screen "15卷绕经验参数" 1280x740, template "模板_调试"
   Group "Group_卷绕经验参数1" at 176,4 size 296x672; FormatPattern 99.99
   Group "Group_卷绕经验参数3" at 808,4 size 296x672; FormatPattern 99.99
   Group "Group_卷绕经验参数2" at 492,4 size 296x672; FormatPattern 99.99
   Button "OBJECT_3" at 176,4 size 80x38; TextOff '支数: / EXIT / 標準糸管１: / 표준보빈1:'
      on Press: SetTag("ST_HMI_Var_HMI_i16_Status_ShaGuan_Select", 1)
   Button "OBJECT_1" at 268,4 size 96x38; TextOff 'f1_n: / EXIT / 標準糸管１: / 표준보빈1:'
      on Press: SetTag("ST_HMI_Var_HMI_i16_Status_ShaGuan_Select", 1)
   Button "OBJECT_2" at 376,4 size 96x38; TextOff 'g1_n: / EXIT / 標準糸管１: / 표준보빈1:'
      on Press: SetTag("ST_HMI_Var_HMI_i16_Status_ShaGuan_Select", 1)
   IOField "IO Field_41" at 176,47 size 80x38; FormatPattern 99.9
      ProcessValue <- "ST_Calculation_Var_1_ZhiShu_ARRAY_JR{3}"
   IOField "IO Field_1" at 268,46 size 96x38; FormatPattern 99.999
      ProcessValue <- "ST_Calculation_Var_1_f1_n_delt_0_n_ARRAY_JR{3}"
   IOField "IO Field_2" at 376,46 size 96x38; FormatPattern 99.999
      ProcessValue <- "ST_Calculation_Var_1_g1_n_delt_0_n_ARRAY_JR{3}"
   IOField "IO Field_3" at 176,89 size 80x38; FormatPattern 99.9
      ProcessValue <- "ST_Calculation_Var_1_ZhiShu_ARRAY_JR{4}"
   IOField "IO Field_4" at 268,88 size 96x38; FormatPattern 99.999
      ProcessValue <- "ST_Calculation_Var_1_f1_n_delt_0_n_ARRAY_JR{4}"
   IOField "IO Field_5" at 376,88 size 96x38; FormatPattern 99.999
      ProcessValue <- "ST_Calculation_Var_1_g1_n_delt_0_n_ARRAY_JR{4}"
   IOField "IO Field_6" at 176,131 size 80x38; FormatPattern 99.9
      ProcessValue <- "ST_Calculation_Var_1_ZhiShu_ARRAY_JR{5}"
   IOField "IO Field_7" at 176,173 size 80x38; FormatPattern 99.9
      ProcessValue <- "ST_Calculation_Var_1_ZhiShu_ARRAY_JR{6}"
   IOField "IO Field_8" at 176,215 size 80x38; FormatPattern 99.9
      ProcessValue <- "ST_Calculation_Var_1_ZhiShu_ARRAY_JR{7}"
   IOField "IO Field_9" at 176,258 size 80x38; FormatPattern 99.9
      ProcessValue <- "ST_Calculation_Var_1_ZhiShu_ARRAY_JR{8}"
   IOField "IO Field_10" at 176,300 size 80x38; FormatPattern 99.9
      ProcessValue <- "ST_Calculation_Var_1_ZhiShu_ARRAY_JR{9}"
   IOField "IO Field_11" at 176,342 size 80x38; FormatPattern 99.9
      ProcessValue <- "ST_Calculation_Var_1_ZhiShu_ARRAY_JR{10}"
   IOField "IO Field_12" at 176,384 size 80x38; FormatPattern 99.9
      ProcessValue <- "ST_Calculation_Var_1_ZhiShu_ARRAY_JR{11}"
   IOField "IO Field_13" at 176,426 size 80x38; FormatPattern 99.9
      ProcessValue <- "ST_Calculation_Var_1_ZhiShu_ARRAY_JR{12}"
   IOField "IO Field_14" at 176,469 size 80x38; FormatPattern 99.9
      ProcessValue <- "ST_Calculation_Var_1_ZhiShu_ARRAY_JR{13}"
   IOField "IO Field_15" at 176,511 size 80x38; FormatPattern 99.9
      ProcessValue <- "ST_Calculation_Var_1_ZhiShu_ARRAY_JR{14}"
   IOField "IO Field_16" at 176,553 size 80x38; FormatPattern 99.9
      ProcessValue <- "ST_Calculation_Var_1_ZhiShu_ARRAY_JR{15}"
   IOField "IO Field_17" at 176,595 size 80x38; FormatPattern 99.9
      ProcessValue <- "ST_Calculation_Var_1_ZhiShu_ARRAY_JR{16}"
   IOField "IO Field_18" at 176,638 size 80x38; FormatPattern 99.9
      ProcessValue <- "ST_Calculation_Var_1_ZhiShu_ARRAY_JR{17}"
   IOField "IO Field_19" at 268,130 size 96x38; FormatPattern 99.999
      ProcessValue <- "ST_Calculation_Var_1_f1_n_delt_0_n_ARRAY_JR{5}"
   IOField "IO Field_20" at 268,172 size 96x38; FormatPattern 99.999
      ProcessValue <- "ST_Calculation_Var_1_f1_n_delt_0_n_ARRAY_JR{6}"
   IOField "IO Field_21" at 268,215 size 96x38; FormatPattern 99.999
      ProcessValue <- "ST_Calculation_Var_1_f1_n_delt_0_n_ARRAY_JR{7}"
   IOField "IO Field_22" at 268,257 size 96x38; FormatPattern 99.999
      ProcessValue <- "ST_Calculation_Var_1_f1_n_delt_0_n_ARRAY_JR{8}"
   IOField "IO Field_23" at 268,299 size 96x38; FormatPattern 99.999
      ProcessValue <- "ST_Calculation_Var_1_f1_n_delt_0_n_ARRAY_JR{9}"
   IOField "IO Field_24" at 268,342 size 96x38; FormatPattern 99.999
      ProcessValue <- "ST_Calculation_Var_1_f1_n_delt_0_n_ARRAY_JR{10}"
   IOField "IO Field_25" at 268,384 size 96x38; FormatPattern 99.999
      ProcessValue <- "ST_Calculation_Var_1_f1_n_delt_0_n_ARRAY_JR{11}"
   IOField "IO Field_26" at 268,426 size 96x38; FormatPattern 99.999
      ProcessValue <- "ST_Calculation_Var_1_f1_n_delt_0_n_ARRAY_JR{12}"
   IOField "IO Field_27" at 268,468 size 96x38; FormatPattern 99.999
      ProcessValue <- "ST_Calculation_Var_1_f1_n_delt_0_n_ARRAY_JR{13}"
   IOField "IO Field_28" at 268,511 size 96x38; FormatPattern 99.999
      ProcessValue <- "ST_Calculation_Var_1_f1_n_delt_0_n_ARRAY_JR{14}"
   IOField "IO Field_29" at 268,553 size 96x38; FormatPattern 99.999
      ProcessValue <- "ST_Calculation_Var_1_f1_n_delt_0_n_ARRAY_JR{15}"
   IOField "IO Field_30" at 268,595 size 96x38; FormatPattern 99.999
      ProcessValue <- "ST_Calculation_Var_1_f1_n_delt_0_n_ARRAY_JR{16}"
   IOField "IO Field_31" at 268,638 size 96x38; FormatPattern 99.999
      ProcessValue <- "ST_Calculation_Var_1_f1_n_delt_0_n_ARRAY_JR{17}"
   IOField "IO Field_32" at 376,130 size 96x38; FormatPattern 99.999
      ProcessValue <- "ST_Calculation_Var_1_g1_n_delt_0_n_ARRAY_JR{5}"
   IOField "IO Field_33" at 376,172 size 96x38; FormatPattern 99.999
      ProcessValue <- "ST_Calculation_Var_1_g1_n_delt_0_n_ARRAY_JR{6}"
   IOField "IO Field_34" at 376,215 size 96x38; FormatPattern 99.999
      ProcessValue <- "ST_Calculation_Var_1_g1_n_delt_0_n_ARRAY_JR{7}"
   IOField "IO Field_35" at 376,257 size 96x38; FormatPattern 99.999
      ProcessValue <- "ST_Calculation_Var_1_g1_n_delt_0_n_ARRAY_JR{8}"
   IOField "IO Field_36" at 376,299 size 96x38; FormatPattern 99.999
      ProcessValue <- "ST_Calculation_Var_1_g1_n_delt_0_n_ARRAY_JR{9}"
   IOField "IO Field_37" at 376,342 size 96x38; FormatPattern 99.999
      ProcessValue <- "ST_Calculation_Var_1_g1_n_delt_0_n_ARRAY_JR{10}"
   IOField "IO Field_38" at 376,384 size 96x38; FormatPattern 99.999
      ProcessValue <- "ST_Calculation_Var_1_g1_n_delt_0_n_ARRAY_JR{11}"
   IOField "IO Field_39" at 376,426 size 96x38; FormatPattern 99.999
      ProcessValue <- "ST_Calculation_Var_1_g1_n_delt_0_n_ARRAY_JR{12}"
   IOField "IO Field_40" at 376,468 size 96x38; FormatPattern 99.999
      ProcessValue <- "ST_Calculation_Var_1_g1_n_delt_0_n_ARRAY_JR{13}"
   IOField "IO Field_42" at 376,511 size 96x38; FormatPattern 99.999
      ProcessValue <- "ST_Calculation_Var_1_g1_n_delt_0_n_ARRAY_JR{14}"
   IOField "IO Field_43" at 376,553 size 96x38; FormatPattern 99.999
      ProcessValue <- "ST_Calculation_Var_1_g1_n_delt_0_n_ARRAY_JR{15}"
   IOField "IO Field_44" at 376,595 size 96x38; FormatPattern 99.999
      ProcessValue <- "ST_Calculation_Var_1_g1_n_delt_0_n_ARRAY_JR{16}"
   IOField "IO Field_45" at 376,638 size 96x38; FormatPattern 99.999
      ProcessValue <- "ST_Calculation_Var_1_g1_n_delt_0_n_ARRAY_JR{17}"
   Button "OBJECT_7" at 808,4 size 80x38; TextOff '支数: / EXIT / 標準糸管１: / 표준보빈1:'
      on Press: SetTag("ST_HMI_Var_HMI_i16_Status_ShaGuan_Select", 1)
   Button "OBJECT_8" at 900,4 size 96x38; TextOff 'f1_n: / EXIT / 標準糸管１: / 표준보빈1:'
      on Press: SetTag("ST_HMI_Var_HMI_i16_Status_ShaGuan_Select", 1)
   Button "OBJECT_9" at 1008,4 size 96x38; TextOff 'g1_n: / EXIT / 標準糸管１: / 표준보빈1:'
      on Press: SetTag("ST_HMI_Var_HMI_i16_Status_ShaGuan_Select", 1)
   IOField "IO Field_91" at 808,47 size 80x38; FormatPattern 99.9
      ProcessValue <- "ST_Calculation_Var_1_ZhiShu_ARRAY_JR{33}"
   IOField "IO Field_92" at 900,46 size 96x38; FormatPattern 99.999
      ProcessValue <- "ST_Calculation_Var_1_f1_n_delt_0_n_ARRAY_JR{33}"
   IOField "IO Field_93" at 1008,46 size 96x38; FormatPattern 99.999
      ProcessValue <- "ST_Calculation_Var_1_g1_n_delt_0_n_ARRAY_JR{33}"
   IOField "IO Field_94" at 808,89 size 80x38; FormatPattern 99.9
      ProcessValue <- "ST_Calculation_Var_1_ZhiShu_ARRAY_JR{34}"
   IOField "IO Field_95" at 900,88 size 96x38; FormatPattern 99.999
      ProcessValue <- "ST_Calculation_Var_1_f1_n_delt_0_n_ARRAY_JR{34}"
   IOField "IO Field_96" at 1008,88 size 96x38; FormatPattern 99.999
      ProcessValue <- "ST_Calculation_Var_1_g1_n_delt_0_n_ARRAY_JR{34}"
   IOField "IO Field_97" at 808,131 size 80x38; FormatPattern 99.9
      ProcessValue <- "ST_Calculation_Var_1_ZhiShu_ARRAY_JR{35}"
   IOField "IO Field_98" at 808,173 size 80x38; FormatPattern 99.9
      ProcessValue <- "ST_Calculation_Var_1_ZhiShu_ARRAY_JR{36}"
   IOField "IO Field_99" at 808,215 size 80x38; FormatPattern 99.9
      ProcessValue <- "ST_Calculation_Var_1_ZhiShu_ARRAY_JR{37}"
   IOField "IO Field_100" at 808,258 size 80x38; FormatPattern 99.9
      ProcessValue <- "ST_Calculation_Var_1_ZhiShu_ARRAY_JR{38}"
   IOField "IO Field_101" at 808,300 size 80x38; FormatPattern 99.9
      ProcessValue <- "ST_Calculation_Var_1_ZhiShu_ARRAY_JR{39}"
   IOField "IO Field_102" at 808,342 size 80x38; FormatPattern 99.9
      ProcessValue <- "ST_Calculation_Var_1_ZhiShu_ARRAY_JR{40}"
   IOField "IO Field_103" at 808,384 size 80x38; FormatPattern 99.9
      ProcessValue <- "ST_Calculation_Var_1_ZhiShu_ARRAY_JR{41}"
   IOField "IO Field_104" at 808,426 size 80x38; FormatPattern 99.9
      ProcessValue <- "ST_Calculation_Var_1_ZhiShu_ARRAY_JR{42}"
   IOField "IO Field_105" at 808,469 size 80x38; FormatPattern 99.9
      ProcessValue <- "ST_Calculation_Var_1_ZhiShu_ARRAY_JR{43}"
   IOField "IO Field_106" at 808,511 size 80x38; FormatPattern 99.9
      ProcessValue <- "ST_Calculation_Var_1_ZhiShu_ARRAY_JR{44}"
   IOField "IO Field_107" at 808,553 size 80x38; FormatPattern 99.9
      ProcessValue <- "ST_Calculation_Var_1_ZhiShu_ARRAY_JR{45}"
   IOField "IO Field_108" at 808,595 size 80x38; FormatPattern 99.9
      ProcessValue <- "ST_Calculation_Var_1_ZhiShu_ARRAY_JR{46}"
   IOField "IO Field_109" at 808,638 size 80x38; FormatPattern 99.9
      ProcessValue <- "ST_Calculation_Var_1_ZhiShu_ARRAY_JR{47}"
   IOField "IO Field_110" at 900,130 size 96x38; FormatPattern 99.999
      ProcessValue <- "ST_Calculation_Var_1_f1_n_delt_0_n_ARRAY_JR{35}"
   IOField "IO Field_111" at 900,172 size 96x38; FormatPattern 99.999
      ProcessValue <- "ST_Calculation_Var_1_f1_n_delt_0_n_ARRAY_JR{36}"
   IOField "IO Field_112" at 900,215 size 96x38; FormatPattern 99.999
      ProcessValue <- "ST_Calculation_Var_1_f1_n_delt_0_n_ARRAY_JR{37}"
   IOField "IO Field_113" at 900,257 size 96x38; FormatPattern 99.999
      ProcessValue <- "ST_Calculation_Var_1_f1_n_delt_0_n_ARRAY_JR{38}"
   IOField "IO Field_114" at 900,299 size 96x38; FormatPattern 99.999
      ProcessValue <- "ST_Calculation_Var_1_f1_n_delt_0_n_ARRAY_JR{39}"
   IOField "IO Field_115" at 900,342 size 96x38; FormatPattern 99.999
      ProcessValue <- "ST_Calculation_Var_1_f1_n_delt_0_n_ARRAY_JR{40}"
   IOField "IO Field_116" at 900,384 size 96x38; FormatPattern 99.999
      ProcessValue <- "ST_Calculation_Var_1_f1_n_delt_0_n_ARRAY_JR{41}"
   IOField "IO Field_117" at 900,426 size 96x38; FormatPattern 99.999
      ProcessValue <- "ST_Calculation_Var_1_f1_n_delt_0_n_ARRAY_JR{42}"
   IOField "IO Field_118" at 900,468 size 96x38; FormatPattern 99.999
      ProcessValue <- "ST_Calculation_Var_1_f1_n_delt_0_n_ARRAY_JR{43}"
   IOField "IO Field_119" at 900,511 size 96x38; FormatPattern 99.999
      ProcessValue <- "ST_Calculation_Var_1_f1_n_delt_0_n_ARRAY_JR{44}"
   IOField "IO Field_120" at 900,553 size 96x38; FormatPattern 99.999
      ProcessValue <- "ST_Calculation_Var_1_f1_n_delt_0_n_ARRAY_JR{45}"
   IOField "IO Field_121" at 900,595 size 96x38; FormatPattern 99.999
      ProcessValue <- "ST_Calculation_Var_1_f1_n_delt_0_n_ARRAY_JR{46}"
   IOField "IO Field_122" at 900,638 size 96x38; FormatPattern 99.999
      ProcessValue <- "ST_Calculation_Var_1_f1_n_delt_0_n_ARRAY_JR{47}"
   IOField "IO Field_123" at 1008,130 size 96x38; FormatPattern 99.999
      ProcessValue <- "ST_Calculation_Var_1_g1_n_delt_0_n_ARRAY_JR{35}"
   IOField "IO Field_124" at 1008,172 size 96x38; FormatPattern 99.999
      ProcessValue <- "ST_Calculation_Var_1_g1_n_delt_0_n_ARRAY_JR{36}"
   IOField "IO Field_125" at 1008,215 size 96x38; FormatPattern 99.999
      ProcessValue <- "ST_Calculation_Var_1_g1_n_delt_0_n_ARRAY_JR{37}"
   IOField "IO Field_126" at 1008,257 size 96x38; FormatPattern 99.999
      ProcessValue <- "ST_Calculation_Var_1_g1_n_delt_0_n_ARRAY_JR{38}"
   IOField "IO Field_127" at 1008,299 size 96x38; FormatPattern 99.999
      ProcessValue <- "ST_Calculation_Var_1_g1_n_delt_0_n_ARRAY_JR{39}"
   IOField "IO Field_128" at 1008,342 size 96x38; FormatPattern 99.999
      ProcessValue <- "ST_Calculation_Var_1_g1_n_delt_0_n_ARRAY_JR{40}"
   IOField "IO Field_129" at 1008,384 size 96x38; FormatPattern 99.999
      ProcessValue <- "ST_Calculation_Var_1_g1_n_delt_0_n_ARRAY_JR{41}"
   IOField "IO Field_130" at 1008,426 size 96x38; FormatPattern 99.999
      ProcessValue <- "ST_Calculation_Var_1_g1_n_delt_0_n_ARRAY_JR{42}"
   IOField "IO Field_131" at 1008,468 size 96x38; FormatPattern 99.999
      ProcessValue <- "ST_Calculation_Var_1_g1_n_delt_0_n_ARRAY_JR{43}"
   IOField "IO Field_132" at 1008,511 size 96x38; FormatPattern 99.999
      ProcessValue <- "ST_Calculation_Var_1_g1_n_delt_0_n_ARRAY_JR{44}"
   IOField "IO Field_133" at 1008,553 size 96x38; FormatPattern 99.999
      ProcessValue <- "ST_Calculation_Var_1_g1_n_delt_0_n_ARRAY_JR{45}"
   IOField "IO Field_134" at 1008,595 size 96x38; FormatPattern 99.999
      ProcessValue <- "ST_Calculation_Var_1_g1_n_delt_0_n_ARRAY_JR{46}"
   IOField "IO Field_135" at 1008,638 size 96x38; FormatPattern 99.999
      ProcessValue <- "ST_Calculation_Var_1_g1_n_delt_0_n_ARRAY_JR{47}"
   Button "OBJECT_4" at 492,4 size 80x38; TextOff '支数: / EXIT / 標準糸管１: / 표준보빈1:'
      on Press: SetTag("ST_HMI_Var_HMI_i16_Status_ShaGuan_Select", 1)
   Button "OBJECT_5" at 584,4 size 96x38; TextOff 'f1_n: / EXIT / 標準糸管１: / 표준보빈1:'
      on Press: SetTag("ST_HMI_Var_HMI_i16_Status_ShaGuan_Select", 1)
   Button "OBJECT_6" at 692,4 size 96x38; TextOff 'g1_n: / EXIT / 標準糸管１: / 표준보빈1:'
      on Press: SetTag("ST_HMI_Var_HMI_i16_Status_ShaGuan_Select", 1)
   IOField "IO Field_46" at 492,47 size 80x38; FormatPattern 99.9
      ProcessValue <- "ST_Calculation_Var_1_ZhiShu_ARRAY_JR{18}"
   IOField "IO Field_47" at 584,46 size 96x38; FormatPattern 99.999
      ProcessValue <- "ST_Calculation_Var_1_f1_n_delt_0_n_ARRAY_JR{18}"
   IOField "IO Field_48" at 692,46 size 96x38; FormatPattern 99.999
      ProcessValue <- "ST_Calculation_Var_1_g1_n_delt_0_n_ARRAY_JR{18}"
   IOField "IO Field_49" at 492,89 size 80x38; FormatPattern 99.9
      ProcessValue <- "ST_Calculation_Var_1_ZhiShu_ARRAY_JR{19}"
   IOField "IO Field_50" at 584,88 size 96x38; FormatPattern 99.999
      ProcessValue <- "ST_Calculation_Var_1_f1_n_delt_0_n_ARRAY_JR{19}"
   IOField "IO Field_51" at 692,88 size 96x38; FormatPattern 99.999
      ProcessValue <- "ST_Calculation_Var_1_g1_n_delt_0_n_ARRAY_JR{19}"
   IOField "IO Field_52" at 492,131 size 80x38; FormatPattern 99.9
      ProcessValue <- "ST_Calculation_Var_1_ZhiShu_ARRAY_JR{20}"
   IOField "IO Field_53" at 492,173 size 80x38; FormatPattern 99.9
      ProcessValue <- "ST_Calculation_Var_1_ZhiShu_ARRAY_JR{21}"
   IOField "IO Field_54" at 492,215 size 80x38; FormatPattern 99.9
      ProcessValue <- "ST_Calculation_Var_1_ZhiShu_ARRAY_JR{22}"
   IOField "IO Field_55" at 492,258 size 80x38; FormatPattern 99.9
      ProcessValue <- "ST_Calculation_Var_1_ZhiShu_ARRAY_JR{23}"
   IOField "IO Field_56" at 492,300 size 80x38; FormatPattern 99.9
      ProcessValue <- "ST_Calculation_Var_1_ZhiShu_ARRAY_JR{24}"
   IOField "IO Field_57" at 492,342 size 80x38; FormatPattern 99.9
      ProcessValue <- "ST_Calculation_Var_1_ZhiShu_ARRAY_JR{25}"
   IOField "IO Field_58" at 492,384 size 80x38; FormatPattern 99.9
      ProcessValue <- "ST_Calculation_Var_1_ZhiShu_ARRAY_JR{26}"
   IOField "IO Field_59" at 492,426 size 80x38; FormatPattern 99.9
      ProcessValue <- "ST_Calculation_Var_1_ZhiShu_ARRAY_JR{27}"
   IOField "IO Field_60" at 492,469 size 80x38; FormatPattern 99.9
      ProcessValue <- "ST_Calculation_Var_1_ZhiShu_ARRAY_JR{28}"
   IOField "IO Field_61" at 492,511 size 80x38; FormatPattern 99.9
      ProcessValue <- "ST_Calculation_Var_1_ZhiShu_ARRAY_JR{29}"
   IOField "IO Field_62" at 492,553 size 80x38; FormatPattern 99.9
      ProcessValue <- "ST_Calculation_Var_1_ZhiShu_ARRAY_JR{30}"
   IOField "IO Field_63" at 492,595 size 80x38; FormatPattern 99.9
      ProcessValue <- "ST_Calculation_Var_1_ZhiShu_ARRAY_JR{31}"
   IOField "IO Field_64" at 492,638 size 80x38; FormatPattern 99.9
      ProcessValue <- "ST_Calculation_Var_1_ZhiShu_ARRAY_JR{32}"
   IOField "IO Field_65" at 584,130 size 96x38; FormatPattern 99.999
      ProcessValue <- "ST_Calculation_Var_1_f1_n_delt_0_n_ARRAY_JR{20}"
   IOField "IO Field_66" at 584,172 size 96x38; FormatPattern 99.999
      ProcessValue <- "ST_Calculation_Var_1_f1_n_delt_0_n_ARRAY_JR{21}"
   IOField "IO Field_67" at 584,215 size 96x38; FormatPattern 99.999
      ProcessValue <- "ST_Calculation_Var_1_f1_n_delt_0_n_ARRAY_JR{22}"
   IOField "IO Field_68" at 584,257 size 96x38; FormatPattern 99.999
      ProcessValue <- "ST_Calculation_Var_1_f1_n_delt_0_n_ARRAY_JR{23}"
   IOField "IO Field_69" at 584,299 size 96x38; FormatPattern 99.999
      ProcessValue <- "ST_Calculation_Var_1_f1_n_delt_0_n_ARRAY_JR{24}"
   IOField "IO Field_70" at 584,342 size 96x38; FormatPattern 99.999
      ProcessValue <- "ST_Calculation_Var_1_f1_n_delt_0_n_ARRAY_JR{25}"
   IOField "IO Field_71" at 584,384 size 96x38; FormatPattern 99.999
      ProcessValue <- "ST_Calculation_Var_1_f1_n_delt_0_n_ARRAY_JR{26}"
   IOField "IO Field_72" at 584,426 size 96x38; FormatPattern 99.999
      ProcessValue <- "ST_Calculation_Var_1_f1_n_delt_0_n_ARRAY_JR{27}"
   IOField "IO Field_73" at 584,468 size 96x38; FormatPattern 99.999
      ProcessValue <- "ST_Calculation_Var_1_f1_n_delt_0_n_ARRAY_JR{28}"
   IOField "IO Field_74" at 584,511 size 96x38; FormatPattern 99.999
      ProcessValue <- "ST_Calculation_Var_1_f1_n_delt_0_n_ARRAY_JR{29}"
   IOField "IO Field_75" at 584,553 size 96x38; FormatPattern 99.999
      ProcessValue <- "ST_Calculation_Var_1_f1_n_delt_0_n_ARRAY_JR{30}"
   IOField "IO Field_76" at 584,595 size 96x38; FormatPattern 99.999
      ProcessValue <- "ST_Calculation_Var_1_f1_n_delt_0_n_ARRAY_JR{31}"
   IOField "IO Field_77" at 584,638 size 96x38; FormatPattern 99.999
      ProcessValue <- "ST_Calculation_Var_1_f1_n_delt_0_n_ARRAY_JR{32}"
   IOField "IO Field_78" at 692,130 size 96x38; FormatPattern 99.999
      ProcessValue <- "ST_Calculation_Var_1_g1_n_delt_0_n_ARRAY_JR{20}"
   IOField "IO Field_79" at 692,172 size 96x38; FormatPattern 99.999
      ProcessValue <- "ST_Calculation_Var_1_g1_n_delt_0_n_ARRAY_JR{21}"
   IOField "IO Field_80" at 692,215 size 96x38; FormatPattern 99.999
      ProcessValue <- "ST_Calculation_Var_1_g1_n_delt_0_n_ARRAY_JR{22}"
   IOField "IO Field_81" at 692,257 size 96x38; FormatPattern 99.999
      ProcessValue <- "ST_Calculation_Var_1_g1_n_delt_0_n_ARRAY_JR{23}"
   IOField "IO Field_82" at 692,299 size 96x38; FormatPattern 99.999
      ProcessValue <- "ST_Calculation_Var_1_g1_n_delt_0_n_ARRAY_JR{24}"
   IOField "IO Field_83" at 692,342 size 96x38; FormatPattern 99.999
      ProcessValue <- "ST_Calculation_Var_1_g1_n_delt_0_n_ARRAY_JR{25}"
   IOField "IO Field_84" at 692,384 size 96x38; FormatPattern 99.999
      ProcessValue <- "ST_Calculation_Var_1_g1_n_delt_0_n_ARRAY_JR{26}"
   IOField "IO Field_85" at 692,426 size 96x38; FormatPattern 99.999
      ProcessValue <- "ST_Calculation_Var_1_g1_n_delt_0_n_ARRAY_JR{27}"
   IOField "IO Field_86" at 692,468 size 96x38; FormatPattern 99.999
      ProcessValue <- "ST_Calculation_Var_1_g1_n_delt_0_n_ARRAY_JR{28}"
   IOField "IO Field_87" at 692,511 size 96x38; FormatPattern 99.999
      ProcessValue <- "ST_Calculation_Var_1_g1_n_delt_0_n_ARRAY_JR{29}"
   IOField "IO Field_88" at 692,553 size 96x38; FormatPattern 99.999
      ProcessValue <- "ST_Calculation_Var_1_g1_n_delt_0_n_ARRAY_JR{30}"
   IOField "IO Field_89" at 692,595 size 96x38; FormatPattern 99.999
      ProcessValue <- "ST_Calculation_Var_1_g1_n_delt_0_n_ARRAY_JR{31}"
   IOField "IO Field_90" at 692,638 size 96x38; FormatPattern 99.999
      ProcessValue <- "ST_Calculation_Var_1_g1_n_delt_0_n_ARRAY_JR{32}"

screen "16机械参数" 1280x740, template "模板_调试"
   GraphicView "图形视图_1" at 395,6 size 437x668; Picture "成形参数_400×600"
   TextField "文本域_1" at 847,6 size 298x260; Text '测绘尺寸: rc0 :成形弓半径 rz0 :张力弓半径 xco :成形弓圆心x坐标 yco :成形弓圆心y坐标 hcz :轴心高度差 H :锭子总高度 Dl :罗拉直径 Hld :锭尖到罗拉顶部的高度 Lld :锭尖到罗拉的距离'
   TextField "文本域_3" at 847,355 size 298x250; Text '绘图后得出的： xzo :张力弓圆心x坐标 yzo :张力弓圆心y坐标 xit_0 :成形弓零位对应的角度 GAM_max :张力弓零位对应的角度 xit_delt_max :成形弓最大行程 gam_delt_max :张力弓最大行程 X_L_0 :罗拉最高点x坐标 Y_L_0 :罗拉最高点y坐标'
   TextField "文本域_2" at 847,270 size 298x80; Text '调整尺寸： hc0 :成形弓零位到锭尖的高度 hz0 :张力弓零位到锭尖的高度'
   TextField "文本域_4" at 143,22 size 145x30; Text '1.rc0'
   TextField "文本域_5" at 143,77 size 145x30; Text '2.rz0'
   TextField "文本域_6" at 143,132 size 145x30; Text '3.xco'
   TextField "文本域_7" at 143,187 size 145x30; Text '4.yco'
   TextField "文本域_8" at 143,242 size 145x30; Text '5.xzo'
   TextField "文本域_9" at 143,297 size 145x30; Text '6.yzo'
   TextField "文本域_10" at 143,352 size 145x30; Text '7.xit_0'
   TextField "文本域_11" at 143,407 size 145x30; Text '8.GAM_max'
   TextField "文本域_12" at 143,462 size 145x30; Text '9.xit_delt_max'
   TextField "文本域_13" at 143,517 size 145x30; Text '10.X_L_0'
   TextField "文本域_14" at 143,572 size 145x30; Text '11.Y_L_0'
   TextField "文本域_15" at 143,628 size 145x30; Text '12.CX_max'
   TextField "文本域_16" at 847,610 size 298x63; Text '设定参数： CX_max :落纱成形最低位置'
   IOField "IO Field_9" at 304,22 size 80x30
      ProcessValue <- "ST_HMI_Var_HMI_rc0"
   IOField "IO Field_1" at 304,77 size 80x30
      ProcessValue <- "ST_HMI_Var_HMI_rz0"
   IOField "IO Field_2" at 304,132 size 80x30
      ProcessValue <- "ST_HMI_Var_HMI_xco"
   IOField "IO Field_3" at 304,187 size 80x30
      ProcessValue <- "ST_HMI_Var_HMI_yco"
   IOField "IO Field_4" at 304,242 size 80x30
      ProcessValue <- "ST_HMI_Var_HMI_xzo"
   IOField "IO Field_5" at 304,297 size 80x30
      ProcessValue <- "ST_HMI_Var_HMI_yzo"
   IOField "IO Field_6" at 304,352 size 80x30
      ProcessValue <- "ST_HMI_Var_HMI_xit_0"
   IOField "IO Field_7" at 304,407 size 80x30
      ProcessValue <- "ST_HMI_Var_HMI_GAM_max"
   IOField "IO Field_8" at 304,462 size 80x30
      ProcessValue <- "ST_HMI_Var_HMI_xit_delt_max"
   IOField "IO Field_10" at 304,517 size 80x30
      ProcessValue <- "ST_HMI_Var_HMI_X_L_0"
   IOField "IO Field_11" at 304,572 size 80x30
      ProcessValue <- "ST_HMI_Var_HMI_Y_L_0"
   IOField "IO Field_12" at 304,628 size 80x30
      ProcessValue <- "ST_HMI_Var_HMI_r64Position_ChengXing_Botton"

Template "模板_根" 1280x740
   Button "template_1_1" at 80,680 size 80x60; TextOn '手动画面'; TextOff '手动操作'; PictureOn "manual_5_500×500_反相"; PictureOff "manual_5_500×500"
      on Release: ActivateScreenByNumber("Picture", 0)
      on Press: SetTag("Picture", 5)
      Appearance <- "Picture"
   Button "template_1_2" at 720,680 size 80x60; TextOn '报警画面'; TextOff '报 警'; PictureOn "emblem_important_1_200×200_反相"; PictureOff "emblem_important_1_200×200"
      on Release: ActivateScreenByNumber("Picture", 0)
      on Press: SetTag("Picture", 6)
      Appearance <- "Picture"
   Button "template_1_5" at 800,680 size 80x60; TextOn '保养提示'; TextOff '保养提示'; PictureOn "baoyang_6_600×600_反相"; PictureOff "baoyang_6_600×600"
      on Release: ActivateScreenByNumber("Picture", 0)
      on Press: SetTag("Picture", 8)
      Appearance <- "Picture"
   Button "template_1_7" at 880,680 size 80x60; TextOn '调试画面'; TextOff '调 试'; Authorization "Operate_4"; PictureOff "kdeconnect-tray_100×100"; PictureOn "kdeconnect-tray_100×100_反相"
      on Release: ActivateScreenByNumber("Picture", 0); function_f23ef4c9()
      on Press: SetTag("Picture", 3)
      Appearance <- "Picture"
   Button "template_1_3" at 0,680 size 80x60; TextOn '手动画面'; TextOff '手动操作'; PictureOff "图形_16"
      on Release: ActivateScreenByNumber("Picture", 0); SetTag("ST_HMI_Var_HMI_i32_ZouChe_ZhanJu_ss_1", 0)
      on Press: function_f23ef4c9(); SetTag("Picture", 1)
      Appearance <- "Picture"
   Button "template_1_4" at 1120,680 size 80x60; TextOff '调 试'; TextOn '调试画面'; Authorization "Operate_4"; PictureOff "System_Shutdown_100×100"; PictureOn "System_Shutdown_反相_100×100"
      on Click: function_f23ef4c9()
      on Release: StopRuntime(0)
   Button "template_1_6" at 1040,680 size 80x60; TextOff 'Text'; TextOn '调试画面'; Authorization "Operate_4"; PictureOff "computer_laptop_100×100"; PictureOn "computer_laptop_100×100_反相"
      on Click: function_f23ef4c9()
      on Release: function_f34a74f3()
   Button "template_1_8" at 960,680 size 80x60; TextOff 'Text'; TextOn '调试画面'; Authorization "Operate_4"; PictureOff "similarartists_amarok_100×100"; PictureOn "similarartists_amarok_100×100_反相"
      on Release: ActivateScreenByNumber("Picture", 0)
      on Press: SetTag("Picture", 7)
      Appearance <- "Picture"
   Button "template_1_23" at 160,680 size 160x60; TextOn '工艺'; TextOff '工艺'; PictureOn "settings_1_32×32_反相"; PictureOff "settings_1_32×32"
      on Release: ActivateScreenByNumber("Picture", 0)
      on Press: SetTag("Picture", 2)
      Appearance <- "Picture"
   TextField "模板_文本域_2" at 320,680 size 400x60; Text '苏州友联纺工装备科技股份有限公司'
   Button "OBJECT_122" at 1200,680 size 80x60; TextOn '响 铃'; TextOff '响 铃 / EXIT'; PictureOn "Gold_bell_100×100_反相"; PictureOff "Gold_bell_100×100"
      on Release: ResetBit("ST_HMI_Var_HMI_bo_XiangLing")
      on Press: SetBit("ST_HMI_Var_HMI_bo_XiangLing")
      Appearance <- "ST_HMI_Var_HMI_bo_XiangLing"

Template "模板_动画" 1280x740
   Bar "棒图_2" at 116,16 size 17x416; MinimumValue -1000; MaximumValue 10500
      ProcessValue <- "ST_HMI_Var_HMI_r64Axis_DingZi_Velocity_real"
   Group "Group_锭子转速" at 163,92 size 84x50
   Group "Group_动画_1" at 160,100 size 1103x448
   Group "Group_捻度" at 163,155 size 98x50
   Button "template_animation_1" at 80,680 size 80x60; TextOn '手动画面'; TextOff '手动操作'; PictureOn "manual_5_500×500_反相"; PictureOff "manual_5_500×500"
      on Release: ActivateScreenByNumber("Picture", 0)
      on Press: SetTag("Picture", 5)
      Appearance <- "Picture"
   Button "template_animation_2" at 720,680 size 80x60; TextOn '报警画面'; TextOff '报 警'; PictureOn "emblem_important_1_200×200_反相"; PictureOff "emblem_important_1_200×200"
      on Release: ActivateScreenByNumber("Picture", 0)
      on Press: SetTag("Picture", 6)
      Appearance <- "Picture"
   Button "template_animation_5" at 800,680 size 80x60; TextOn '保养提示'; TextOff '保养提示'; PictureOn "baoyang_6_600×600_反相"; PictureOff "baoyang_6_600×600"
      on Release: ActivateScreenByNumber("Picture", 0)
      on Press: SetTag("Picture", 8)
      Appearance <- "Picture"
   Button "template_animation_7" at 880,680 size 80x60; TextOn '调试画面'; TextOff '调 试'; Authorization "Operate_4"; PictureOff "kdeconnect-tray_100×100"; PictureOn "kdeconnect-tray_100×100_反相"
      on Release: ActivateScreenByNumber("Picture", 0); function_f23ef4c9()
      on Press: SetTag("Picture", 3)
      Appearance <- "Picture"
   Button "template_animation_3" at 0,680 size 80x60; TextOn '手动画面'; TextOff '手动操作'; PictureOff "图形_16"
      on Release: ActivateScreenByNumber("Picture", 0); SetTag("ST_HMI_Var_HMI_i32_ZouChe_ZhanJu_ss_1", 0)
      on Press: function_f23ef4c9(); SetTag("Picture", 1)
      Appearance <- "Picture"
   Button "template_animation_4" at 1120,680 size 80x60; TextOff '调 试'; TextOn '调试画面'; PictureOn "System_Shutdown_反相_100×100"; PictureOff "System_Shutdown_100×100"; Authorization "Operate_4"
      on Click: function_f23ef4c9()
      on Release: StopRuntime(0)
   Button "template_animation_6" at 1040,680 size 80x60; TextOff 'Text'; TextOn '调试画面'; PictureOn "computer_laptop_100×100_反相"; PictureOff "computer_laptop_100×100"; Authorization "Operate_4"
      on Click: function_f23ef4c9()
      on Release: function_f34a74f3()
   Button "template_animation_8" at 960,680 size 80x60; TextOff 'Text'; TextOn '调试画面'; PictureOn "similarartists_amarok_100×100_反相"; PictureOff "similarartists_amarok_100×100"; Authorization "Operate_4"
      on Release: ActivateScreenByNumber("Picture", 0)
      on Press: SetTag("Picture", 7)
      Appearance <- "Picture"
   Rectangle "模板_矩形_2" at 559,499 size 552x50
      Visibility <- "ST_Main_Var_g_bo_Automatic_Running_Status"
   Button "template_animation_23" at 160,680 size 160x60; TextOn '工艺'; TextOff '工艺'; PictureOn "settings_1_32×32_反相"; PictureOff "settings_1_32×32"
      on Release: ActivateScreenByNumber("Picture", 0)
      on Press: SetTag("Picture", 2)
      Appearance <- "Picture"
   TextField "模板_文本域_2" at 320,680 size 400x60; Text '苏州友联纺工装备科技股份有限公司'
   IOField "IO Field_57" at 163,92 size 51x25; FormatPattern 99999
      ProcessValue <- "ST_HMI_Var_HMI_r64Axis_DingZi_Velocity_real"
   TextField "文本域_9" at 213,92 size 34x25; Text '/'
   IOField "IO Field_56" at 163,117 size 51x25; FormatPattern 99999
      ProcessValue <- "ST_HMI_Var_HMI_r64Axis_DingZi_Velocity_object"
   TextField "文本域_10" at 213,117 size 34x25; Text 'rpm'
   Group "Group_纱穗" at 11,16 size 78x416
   Polygon "多边形_195" at 11,122 size 78x280
      Visibility <- "VBS_hengsi_status1"
   Polygon "多边形_196" at 11,207 size 78x195
      Visibility <- "VBS_hengsi_status1"
   Polygon "多边形_264" at 32,301 size 38x101
      Visibility <- "VBS_hengsi_status0"
   Polygon "多边形_265" at 36,312 size 29x90
      Visibility <- "VBS_hengsi_status0"
   Polygon "多边形_198" at 11,116 size 78x286
      Visibility <- "VBS_hengsi_status1"
   Polygon "多边形_199" at 11,201 size 78x200
      Visibility <- "VBS_hengsi_status1"
   Polygon "多边形_266" at 29,293 size 42x107
      Visibility <- "VBS_hengsi_status0"
   Polygon "多边形_201" at 11,112 size 78x289
      Visibility <- "VBS_hengsi_status1"
   Polygon "多边形_202" at 11,198 size 78x204
      Visibility <- "VBS_hengsi_status1"
   Polygon "多边形_267" at 27,285 size 47x117
      Visibility <- "VBS_hengsi_status0"
   Polygon "多边形_204" at 11,110 size 78x292
      Visibility <- "VBS_hengsi_status1"
   Polygon "多边形_205" at 11,193 size 78x209
      Visibility <- "VBS_hengsi_status1"
   Polygon "多边形_268" at 25,278 size 50x124
      Visibility <- "VBS_hengsi_status0"
   Polygon "多边形_207" at 11,106 size 78x296
      Visibility <- "VBS_hengsi_status1"
   Polygon "多边形_208" at 11,190 size 78x211
      Visibility <- "VBS_hengsi_status1"
   Polygon "多边形_269" at 24,273 size 52x128
      Visibility <- "VBS_hengsi_status0"
   Polygon "多边形_210" at 11,101 size 78x301
      Visibility <- "VBS_hengsi_status0"
   Polygon "多边形_211" at 11,187 size 78x215
      Visibility <- "VBS_hengsi_status1"
   Polygon "多边形_270" at 24,266 size 52x135
      Visibility <- "VBS_hengsi_status0"
   Polygon "多边形_213" at 11,97 size 78x304
      Visibility <- "VBS_hengsi_status1"
   Polygon "多边形_214" at 11,183 size 78x218
      Visibility <- "VBS_hengsi_status1"
   Polygon "多边形_271" at 23,261 size 55x140
      Visibility <- "VBS_hengsi_status0"
   Polygon "多边形_216" at 11,92 size 78x309
      Visibility <- "VBS_hengsi_status1"
   Polygon "多边形_217" at 11,178 size 78x224
      Visibility <- "VBS_hengsi_status1"
   Polygon "多边形_272" at 23,258 size 55x144
      Visibility <- "VBS_hengsi_status0"
   Polygon "多边形_219" at 11,89 size 78x313
      Visibility <- "VBS_hengsi_status1"
   Polygon "多边形_220" at 11,175 size 78x227
      Visibility <- "VBS_hengsi_status1"
   Polygon "多边形_273" at 21,255 size 57x146
      Visibility <- "VBS_hengsi_status0"
   Polygon "多边形_222" at 11,86 size 78x315
      Visibility <- "VBS_hengsi_status1"
   Polygon "多边形_223" at 11,172 size 78x230
      Visibility <- "VBS_hengsi_status1"
   Polygon "多边形_274" at 21,253 size 57x148
      Visibility <- "VBS_hengsi_status0"
   Polygon "多边形_225" at 11,83 size 78x319
      Visibility <- "VBS_hengsi_status1"
   Polygon "多边形_226" at 11,169 size 78x233
      Visibility <- "VBS_hengsi_status1"
   Polygon "多边形_275" at 21,250 size 59x152
      Visibility <- "VBS_hengsi_status0"
   Polygon "多边形_228" at 11,78 size 78x324
      Visibility <- "VBS_hengsi_status1"
   Polygon "多边形_229" at 11,163 size 78x238
      Visibility <- "VBS_hengsi_status1"
   Polygon "多边形_276" at 21,247 size 59x155
      Visibility <- "VBS_hengsi_status0"
   Polygon "多边形_231" at 11,74 size 78x328
      Visibility <- "VBS_hengsi_status1"
   Polygon "多边形_232" at 11,160 size 78x242
      Visibility <- "VBS_hengsi_status1"
   Polygon "多边形_277" at 19,243 size 61x159
      Visibility <- "VBS_hengsi_status0"
   Polygon "多边形_234" at 11,69 size 78x333
      Visibility <- "VBS_hengsi_status1"
   Polygon "多边形_235" at 11,155 size 78x247
      Visibility <- "VBS_hengsi_status1"
   Polygon "多边形_278" at 17,243 size 64x159
      Visibility <- "VBS_hengsi_status0"
   Polygon "多边形_237" at 11,68 size 78x334
      Visibility <- "VBS_hengsi_status1"
   Polygon "多边形_238" at 11,151 size 78x250
      Visibility <- "VBS_hengsi_status1"
   Polygon "多边形_279" at 17,240 size 64x162
      Visibility <- "VBS_hengsi_status0"
   Polygon "多边形_240" at 11,63 size 78x339
      Visibility <- "VBS_hengsi_status1"
   Polygon "多边形_241" at 11,149 size 78x253
      Visibility <- "VBS_hengsi_status1"
   Polygon "多边形_280" at 16,236 size 67x166
      Visibility <- "VBS_hengsi_status0"
   Polygon "多边形_243" at 11,59 size 78x342
      Visibility <- "VBS_hengsi_status1"
   Polygon "多边形_244" at 11,145 size 78x257
      Visibility <- "VBS_hengsi_status1"
   Polygon "多边形_281" at 16,234 size 67x167
      Visibility <- "VBS_hengsi_status0"
   Polygon "多边形_246" at 11,54 size 78x348
      Visibility <- "VBS_hengsi_status1"
   Polygon "多边形_247" at 11,140 size 78x262
      Visibility <- "VBS_hengsi_status1"
   Polygon "多边形_282" at 15,232 size 68x170
      Visibility <- "VBS_hengsi_status0"
   Polygon "多边形_249" at 11,51 size 78x351
      Visibility <- "VBS_hengsi_status1"
   Polygon "多边形_250" at 11,136 size 78x265
      Visibility <- "VBS_hengsi_status1"
   Polygon "多边形_283" at 15,228 size 68x173
      Visibility <- "VBS_hengsi_status0"
   Polygon "多边形_252" at 11,47 size 78x354
      Visibility <- "VBS_hengsi_status1"
   Polygon "多边形_253" at 11,131 size 78x270
      Visibility <- "VBS_hengsi_status1"
   Polygon "多边形_284" at 14,225 size 72x177
      Visibility <- "VBS_hengsi_status0"
   Polygon "多边形_255" at 11,45 size 78x357
      Visibility <- "VBS_hengsi_status1"
   Polygon "多边形_256" at 11,130 size 78x271
      Visibility <- "VBS_hengsi_status1"
   Polygon "多边形_285" at 14,221 size 72x180
      Visibility <- "VBS_hengsi_status0"
   Polygon "多边形_258" at 11,125 size 78x276
      Visibility <- "VBS_hengsi_status1"
   Polygon "多边形_286" at 13,218 size 74x184
      Visibility <- "VBS_hengsi_status0"
   Polygon "多边形_287" at 13,214 size 74x187
      Visibility <- "VBS_hengsi_status0"
   Polygon "多边形_288" at 11,214 size 76x188
      Visibility <- "VBS_hengsi_status0"
   Polygon "多边形_289" at 11,208 size 78x193
      Visibility <- "VBS_hengsi_status0"
   Button "OBJECT_122" at 1200,680 size 80x60; TextOn '响 铃'; TextOff '响 铃 / EXIT'; PictureOn "Gold_bell_100×100_反相"; PictureOff "Gold_bell_100×100"
      on Release: ResetBit("ST_HMI_Var_HMI_bo_XiangLing")
      on Press: SetBit("ST_HMI_Var_HMI_bo_XiangLing")
      Appearance <- "ST_HMI_Var_HMI_bo_XiangLing"
   Line "line_3" at 376,225 size 666x17
      Visibility <- "ST_HMI_Var_HMI_r64Axis_1_ZhangLi_Position_JuanRao_real2"
   Line "line_4" at 376,225 size 666x15
      Visibility <- "ST_HMI_Var_HMI_r64Axis_1_ZhangLi_Position_JuanRao_real2"
   Line "line_5" at 378,229 size 664x12
      Visibility <- "ST_HMI_Var_HMI_r64Axis_1_ZhangLi_Position_JuanRao_real2"
   Line "line_6" at 379,232 size 662x9
      Visibility <- "ST_HMI_Var_HMI_r64Axis_1_ZhangLi_Position_JuanRao_real2"
   Line "line_7" at 381,236 size 660x5
      Visibility <- "ST_HMI_Var_HMI_r64Axis_1_ZhangLi_Position_JuanRao_real2"
   Line "line_8" at 381,239 size 660x2
      Visibility <- "ST_HMI_Var_HMI_r64Axis_1_ZhangLi_Position_JuanRao_real2"
   Line "line_12" at 381,241 size 660x5
      Visibility <- "ST_HMI_Var_HMI_r64Axis_1_ZhangLi_Position_JuanRao_real2"
   Line "line_13" at 383,241 size 659x9
      Visibility <- "ST_HMI_Var_HMI_r64Axis_1_ZhangLi_Position_JuanRao_real2"
   Line "line_14" at 383,241 size 659x12
      Visibility <- "ST_HMI_Var_HMI_r64Axis_1_ZhangLi_Position_JuanRao_real2"
   Line "line_27" at 345,239 size 699x17
      Visibility <- "ST_HMI_Var_HMI_r64Axis_1_ZhangLi_Position_JuanRao_real2"
   Line "line_1" at 345,239 size 697x17
      Visibility <- "ST_Main_Var_g_i16_Automatic_Status"
   Group "Group_8" at 387,320 size 876x151
   Group "Group_罗拉位置" at 398,158 size 82x49
      DirectMovement <- "ST_HMI_Var_HMI_r64Axis_ZouChe_Position_real2"
   Group "Group_总牵伸" at 398,109 size 116x25
      DirectMovement <- "ST_HMI_Var_HMI_r64Axis_ZouChe_Position_real2"
   Button "OBJECT_112" at 560,500 size 110x48; TextOff '出车 / EXIT'; Authorization "User administration"
      on Press: SetTag("ST_Main_Var_g_i16_Automatic_Selected", 8); function_f23ef4c9()
      Appearance <- "ST_Main_Var_g_i16_Automatic_Selected"
      Visibility <- "ST_Main_Var_g_i16_Mode_Enabled"
   Button "OBJECT_113" at 670,500 size 110x48; TextOff '出车到 / EXIT'; Authorization "User administration"
      on Press: SetTag("ST_Main_Var_g_i16_Automatic_Selected", 16); function_f23ef4c9()
      Appearance <- "ST_Main_Var_g_i16_Automatic_Selected"
      Visibility <- "ST_Main_Var_g_i16_Mode_Enabled"
   Button "OBJECT_114" at 780,500 size 110x48; TextOff '退绕 / EXIT'; Authorization "User administration"
      on Press: SetTag("ST_Main_Var_g_i16_Automatic_Selected", 32); function_f23ef4c9()
      Appearance <- "ST_Main_Var_g_i16_Automatic_Selected"
      Visibility <- "ST_Main_Var_g_i16_Mode_Enabled"
   Button "OBJECT_115" at 890,500 size 110x48; TextOff '卷绕 / EXIT'; Authorization "User administration"
      on Press: SetTag("ST_Main_Var_g_i16_Automatic_Selected", 64); function_f23ef4c9()
      Appearance <- "ST_Main_Var_g_i16_Automatic_Selected"
      Visibility <- "ST_Main_Var_g_i16_Mode_Enabled"
   Button "OBJECT_116" at 1000,500 size 110x48; TextOff '存绕 / EXIT'; Authorization "User administration"
      on Press: SetTag("ST_Main_Var_g_i16_Automatic_Selected", 128); function_f23ef4c9()
      Appearance <- "ST_Main_Var_g_i16_Automatic_Selected"
      Visibility <- "ST_Main_Var_g_i16_Mode_Enabled"
   TextField "文本域_13" at 460,378 size 51x28; Text 'sec'
   TextField "文本域_14" at 576,378 size 64x28; Text 'm/min'
   IOField "IO Field_81" at 389,381 size 72x28; FormatPattern 999.99
      ProcessValue <- "ST_Main_Var_g_r64_Time_Once"
   IOField "IO Field_82" at 505,381 size 72x28; FormatPattern 999.99
      ProcessValue <- "ST_Main_Var_g_r64_Length_One_Minute"
   TextField "模板_文本域_1" at 161,465 size 77x25; Text '友联装备'
   Group "Group_1" at 299,226 size 76x206
   Group "Group_5" at 202,225 size 173x216
   Group "Group" at 278,256 size 73x216
   Group "Group_11" at 162,225 size 228x110
   Group "Group_6" at 160,296 size 75x46
   Group "Group_12" at 1053,375 size 118x39
   Rectangle "矩形_3" at 404,212 size 191x69
      DirectMovement <- "ST_HMI_Var_HMI_r64Axis_ZouChe_Position_real2"
   Rectangle "矩形_5" at 581,212 size 185x69
      DirectMovement <- "ST_HMI_Var_HMI_r64Axis_ZouChe_Position_real2"
   Rectangle "矩形_7" at 766,212 size 185x69
      DirectMovement <- "ST_HMI_Var_HMI_r64Axis_ZouChe_Position_real2"
   Rectangle "矩形_8" at 951,212 size 185x69
      DirectMovement <- "ST_HMI_Var_HMI_r64Axis_ZouChe_Position_real2"
   Group "Group_车架_V1_001" at 398,100 size 195x272
      DirectMovement <- "ST_HMI_Var_HMI_r64Axis_ZouChe_Position_real2"
   Group "Group_走车位置" at 420,323 size 158x25
      DirectMovement <- "ST_HMI_Var_HMI_r64Axis_ZouChe_Position_real2"
   Group "Group_成形&张力" at 163,221 size 90x48
   IOField "IO Field_66" at 398,158 size 60x25; FormatPattern 9999.9
      ProcessValue <- "Axis_LuoLa_positioningState_commandPosition"
   IOField "IO Field_65" at 398,182 size 60x25; FormatPattern 9999.9
      ProcessValue <- "ST_Main_Var_g_r64Axis_LuoLa_Position"
   TextField "文本域_4" at 458,158 size 22x25; Text '/'
   TextField "文本域_5" at 458,182 size 22x25; Text 'mm'
   IOField "IO Field_60" at 398,109 size 51x25; FormatPattern 9.999
      ProcessValue <- "ST_HMI_Var_HMI_r64QianShen_All_real"
   TextField "文本域_8" at 449,109 size 16x25; Text '/'
   IOField "IO Field_59" at 463,109 size 51x25; FormatPattern 9.999
      ProcessValue <- "ST_HMI_Var_HMI_r64QianShen_All_object"
   Polyline "折线_1" at 302,226 size 73x198
      Visibility <- "ST_HMI_Var_HMI_r64Axis_ChengXing_Position_real2"
   Polyline "折线_25" at 315,226 size 60x154
      Visibility <- "ST_HMI_Var_HMI_r64Axis_ChengXing_Position_real2"
   Polyline "折线_37" at 331,226 size 44x101
      Visibility <- "ST_HMI_Var_HMI_r64Axis_ChengXing_Position_real2"
   Polyline "折线_45" at 345,226 size 30x49
      Visibility <- "ST_HMI_Var_HMI_r64Axis_ChengXing_Position_real2"
   Polyline "折线_46" at 307,226 size 68x200
      Visibility <- "ST_HMI_Var_HMI_r64Axis_ChengXing_Position_real2"
   Polyline "折线_50" at 315,226 size 60x155
      Visibility <- "ST_HMI_Var_HMI_r64Axis_ChengXing_Position_real2"
   Polyline "折线_51" at 331,226 size 44x105
      Visibility <- "ST_HMI_Var_HMI_r64Axis_ChengXing_Position_real2"
   Polyline "折线_57" at 345,226 size 30x52
      Visibility <- "ST_HMI_Var_HMI_r64Axis_ChengXing_Position_real2"
   Polyline "折线_68" at 307,226 size 68x202
      Visibility <- "ST_HMI_Var_HMI_r64Axis_ChengXing_Position_real2"
   Polyline "折线_71" at 315,226 size 60x158
      Visibility <- "ST_HMI_Var_HMI_r64Axis_ChengXing_Position_real2"
   Polyline "折线_72" at 331,226 size 44x106
      Visibility <- "ST_HMI_Var_HMI_r64Axis_ChengXing_Position_real2"
   Polyline "折线_77" at 345,226 size 30x54
      Visibility <- "ST_HMI_Var_HMI_r64Axis_ChengXing_Position_real2"
   Polyline "折线_78" at 302,226 size 73x203
      Visibility <- "ST_HMI_Var_HMI_r64Axis_ChengXing_Position_real2"
   Polyline "折线_79" at 312,226 size 63x161
      Visibility <- "ST_HMI_Var_HMI_r64Axis_ChengXing_Position_real2"
   Polyline "折线_80" at 326,226 size 49x109
      Visibility <- "ST_HMI_Var_HMI_r64Axis_ChengXing_Position_real2"
   Polyline "折线_81" at 340,226 size 35x57
      Visibility <- "ST_HMI_Var_HMI_r64Axis_ChengXing_Position_real2"
   Polyline "折线_82" at 299,226 size 76x206
      Visibility <- "ST_HMI_Var_HMI_r64Axis_ChengXing_Position_real2"
   Polyline "折线_83" at 340,226 size 35x59
      Visibility <- "ST_HMI_Var_HMI_r64Axis_ChengXing_Position_real2"
   Polyline "折线_84" at 331,226 size 44x112
      Visibility <- "ST_HMI_Var_HMI_r64Axis_ChengXing_Position_real2"
   Polyline "折线_85" at 312,226 size 63x163
      Visibility <- "ST_HMI_Var_HMI_r64Axis_ChengXing_Position_real2"
   Polyline "折线_86" at 312,226 size 63x165
      Visibility <- "ST_HMI_Var_HMI_r64Axis_ChengXing_Position_real2"
   Polyline "折线_87" at 322,226 size 53x114
      Visibility <- "ST_HMI_Var_HMI_r64Axis_ChengXing_Position_real2"
   Polyline "折线_88" at 340,226 size 35x62
      Visibility <- "ST_HMI_Var_HMI_r64Axis_ChengXing_Position_real2"
   Polyline "折线_89" at 315,226 size 60x167
      Visibility <- "ST_HMI_Var_HMI_r64Axis_ChengXing_Position_real2"
   Polyline "折线_90" at 321,226 size 54x117
      Visibility <- "ST_HMI_Var_HMI_r64Axis_ChengXing_Position_real2"
   Polyline "折线_91" at 340,226 size 35x64
      Visibility <- "ST_HMI_Var_HMI_r64Axis_ChengXing_Position_real2"
   Polyline "折线_92" at 312,226 size 63x170
      Visibility <- "ST_HMI_Var_HMI_r64Axis_ChengXing_Position_real2"
   Polyline "折线_93" at 326,226 size 49x120
      Visibility <- "ST_HMI_Var_HMI_r64Axis_ChengXing_Position_real2"
   Polyline "折线_94" at 340,226 size 35x67
      Visibility <- "ST_HMI_Var_HMI_r64Axis_ChengXing_Position_real2"
   Polyline "折线_95" at 312,226 size 63x171
      Visibility <- "ST_HMI_Var_HMI_r64Axis_ChengXing_Position_real2"
   Polyline "折线_96" at 321,226 size 54x123
      Visibility <- "ST_HMI_Var_HMI_r64Axis_ChengXing_Position_real2"
   Polyline "折线_97" at 334,226 size 41x70
      Visibility <- "ST_HMI_Var_HMI_r64Axis_ChengXing_Position_real2"
   Polyline "折线_98" at 312,226 size 63x173
      Visibility <- "ST_HMI_Var_HMI_r64Axis_ChengXing_Position_real2"
   Polyline "折线_99" at 326,226 size 49x125
      Visibility <- "ST_HMI_Var_HMI_r64Axis_ChengXing_Position_real2"
   Polyline "折线_100" at 340,226 size 35x72
      Visibility <- "ST_HMI_Var_HMI_r64Axis_ChengXing_Position_real2"
   Polyline "折线_101" at 305,226 size 70x176
      Visibility <- "ST_HMI_Var_HMI_r64Axis_ChengXing_Position_real2"
   Polyline "折线_102" at 321,226 size 54x128
      Visibility <- "ST_HMI_Var_HMI_r64Axis_ChengXing_Position_real2"
   Polyline "折线_103" at 334,226 size 41x75
      Visibility <- "ST_HMI_Var_HMI_r64Axis_ChengXing_Position_real2"
   Polyline "折线_104" at 307,226 size 68x178
      Visibility <- "ST_HMI_Var_HMI_r64Axis_ChengXing_Position_real2"
   Polyline "折线_105" at 334,226 size 41x78
      Visibility <- "ST_HMI_Var_HMI_r64Axis_ChengXing_Position_real2"
   Polyline "折线_106" at 326,226 size 49x131
      Visibility <- "ST_HMI_Var_HMI_r64Axis_ChengXing_Position_real2"
   Polyline "折线_107" at 307,226 size 68x181
      Visibility <- "ST_HMI_Var_HMI_r64Axis_ChengXing_Position_real2"
   Polyline "折线_108" at 321,226 size 54x134
      Visibility <- "ST_HMI_Var_HMI_r64Axis_ChengXing_Position_real2"
   Polyline "折线_109" at 334,226 size 41x81
      Visibility <- "ST_HMI_Var_HMI_r64Axis_ChengXing_Position_real2"
   Polyline "折线_110" at 307,226 size 68x183
      Visibility <- "ST_HMI_Var_HMI_r64Axis_ChengXing_Position_real2"
   Polyline "折线_111" at 334,226 size 41x82
      Visibility <- "ST_HMI_Var_HMI_r64Axis_ChengXing_Position_real2"
   Polyline "折线_112" at 321,226 size 54x136
      Visibility <- "ST_HMI_Var_HMI_r64Axis_ChengXing_Position_real2"
   Polyline "折线_113" at 308,226 size 67x185
      Visibility <- "ST_HMI_Var_HMI_r64Axis_ChengXing_Position_real2"
   Polyline "折线_114" at 321,226 size 54x138
      Visibility <- "ST_HMI_Var_HMI_r64Axis_ChengXing_Position_real2"
   Polyline "折线_115" at 334,226 size 41x86
      Visibility <- "ST_HMI_Var_HMI_r64Axis_ChengXing_Position_real2"
   Polyline "折线_116" at 315,226 size 60x142
      Visibility <- "ST_HMI_Var_HMI_r64Axis_ChengXing_Position_real2"
   Polyline "折线_117" at 307,226 size 68x188
      Visibility <- "ST_HMI_Var_HMI_r64Axis_ChengXing_Position_real2"
   Polyline "折线_118" at 334,226 size 41x89
      Visibility <- "ST_HMI_Var_HMI_r64Axis_ChengXing_Position_real2"
   Polyline "折线_119" at 307,226 size 68x190
      Visibility <- "ST_HMI_Var_HMI_r64Axis_ChengXing_Position_real2"
   Polyline "折线_120" at 334,226 size 41x91
      Visibility <- "ST_HMI_Var_HMI_r64Axis_ChengXing_Position_real2"
   Polyline "折线_121" at 321,226 size 54x144
      Visibility <- "ST_HMI_Var_HMI_r64Axis_ChengXing_Position_real2"
   Polyline "折线_122" at 307,226 size 68x191
      Visibility <- "ST_HMI_Var_HMI_r64Axis_ChengXing_Position_real2"
   Polyline "折线_123" at 315,226 size 60x146
      Visibility <- "ST_HMI_Var_HMI_r64Axis_ChengXing_Position_real2"
   Polyline "折线_124" at 331,226 size 44x94
      Visibility <- "ST_HMI_Var_HMI_r64Axis_ChengXing_Position_real2"
   Polyline "折线_125" at 303,226 size 72x193
      Visibility <- "ST_HMI_Var_HMI_r64Axis_ChengXing_Position_real2"
   Polyline "折线_126" at 327,226 size 48x96
      Visibility <- "ST_HMI_Var_HMI_r64Axis_ChengXing_Position_real2"
   Polyline "折线_127" at 315,226 size 60x148
      Visibility <- "ST_HMI_Var_HMI_r64Axis_ChengXing_Position_real2"
   Polyline "折线_128" at 307,226 size 68x196
      Visibility <- "ST_HMI_Var_HMI_r64Axis_ChengXing_Position_real2"
   Polyline "折线_129" at 331,226 size 44x99
      Visibility <- "ST_HMI_Var_HMI_r64Axis_ChengXing_Position_real2"
   Polyline "折线_130" at 315,226 size 60x151
      Visibility <- "ST_HMI_Var_HMI_r64Axis_ChengXing_Position_real2"
   Group "Group_3" at 202,225 size 173x216
   Group "Group_4" at 202,225 size 173x216
   Line "线_1" at 219,318 size 156x8
      Visibility <- "ST_HMI_Var_HMI_r64Axis_ChengXing_Position_real2"
   Line "线_2" at 219,318 size 144x58
      Visibility <- "ST_HMI_Var_HMI_r64Axis_ChengXing_Position_real2"